REGION Network 10: Concatenadora 10
   RUNG wire#powerrail
      Contact( "EstadosCmpALTA-MTA"._6s1 )
      I_Contact( "CompALTA-MTA".ReqMch6 )
      wire#w1
      Contact( "DB-CompAltaDatos".Aut6 )
      Coil( "Concatenadoras"._6c10 )
   END_RUNG
   RUNG wire#powerrail
      Contact( "EstadosCmpALTA-MTA"._6s9 )
      I_Contact( "CompALTA-MTA".ReqMch6 )
   END_RUNG wire#w1
   RUNG wire#powerrail
      Contact( "EstadosCmpALTA-MTA"._6s3 )
      I_Contact( "DB-CompAltaDatos".PanMchCmp6 )
   END_RUNG wire#w1
   // the same network as SCL:
   "Concatenadoras"._6c10 := (("EstadosCmpALTA-MTA"._6s1 AND NOT "CompALTA-MTA".ReqMch6) OR ("EstadosCmpALTA-MTA"._6s9 AND NOT "CompALTA-MTA".ReqMch6) OR ("EstadosCmpALTA-MTA"._6s3 AND NOT "DB-CompAltaDatos".PanMchCmp6)) AND "DB-CompAltaDatos".Aut6;
END_REGION

REGION Network 11: Concatenadora 4
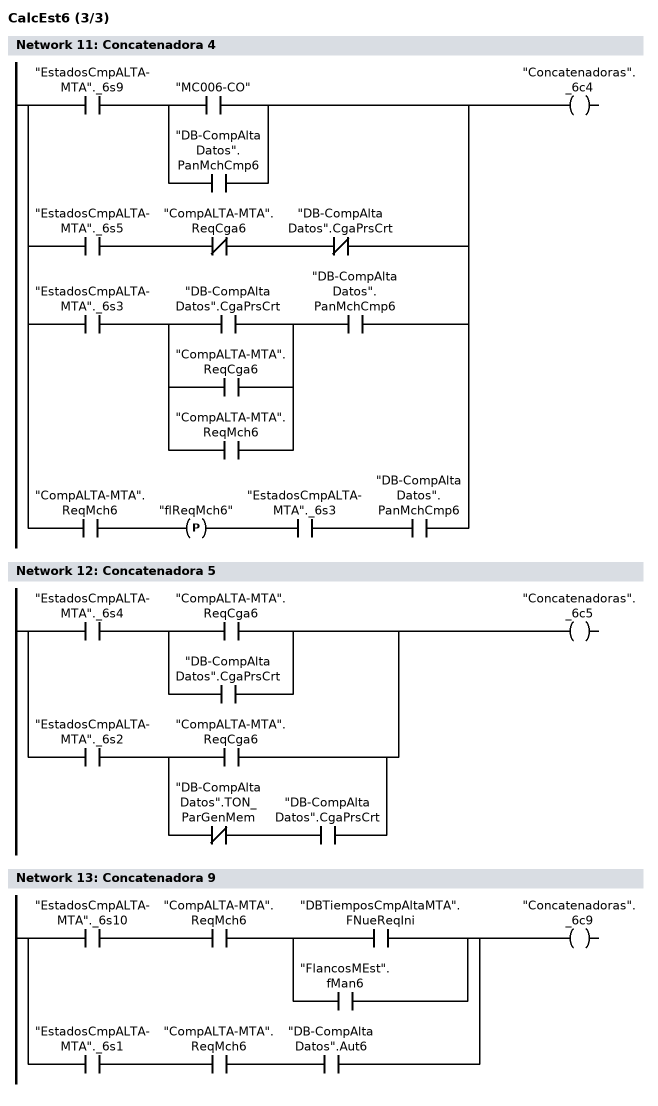
   RUNG wire#powerrail
      Contact( "EstadosCmpALTA-MTA"._6s9 )
      wire#w1
      Contact( "MC006-CO" )
      wire#w2
      Coil( "Concatenadoras"._6c4 )
   END_RUNG
   RUNG wire#w1
      Contact( "DB-CompAltaDatos".PanMchCmp6 )
   END_RUNG wire#w2
   RUNG wire#powerrail
      Contact( "EstadosCmpALTA-MTA"._6s5 )
      I_Contact( "CompALTA-MTA".ReqCga6 )
      I_Contact( "DB-CompAltaDatos".CgaPrsCrt )
   END_RUNG wire#w2
   RUNG wire#powerrail
      Contact( "EstadosCmpALTA-MTA"._6s3 )
      wire#w3
      Contact( "DB-CompAltaDatos".CgaPrsCrt )
      wire#w4
      Contact( "DB-CompAltaDatos".PanMchCmp6 )
   END_RUNG wire#w2
   RUNG wire#w3
      Contact( "CompALTA-MTA".ReqCga6 )
   END_RUNG wire#w4
   RUNG wire#w3
      Contact( "CompALTA-MTA".ReqMch6 )
   END_RUNG wire#w4
   RUNG wire#powerrail
      Contact( "CompALTA-MTA".ReqMch6 )
      P_Trig( "flReqMch6" )
      Contact( "EstadosCmpALTA-MTA"._6s3 )
      Contact( "DB-CompAltaDatos".PanMchCmp6 )
   END_RUNG wire#w2
   // the same network as SCL:
   #_w1 := "CompALTA-MTA".ReqMch6 AND NOT "flReqMch6";   // rising edge
   "flReqMch6" := "CompALTA-MTA".ReqMch6;
   "Concatenadoras"._6c4 := ("EstadosCmpALTA-MTA"._6s9 AND ("MC006-CO" OR "DB-CompAltaDatos".PanMchCmp6)) OR ("EstadosCmpALTA-MTA"._6s5 AND NOT "CompALTA-MTA".ReqCga6 AND NOT "DB-CompAltaDatos".CgaPrsCrt) OR ("EstadosCmpALTA-MTA"._6s3 AND ("DB-CompAltaDatos".CgaPrsCrt OR "CompALTA-MTA".ReqCga6 OR "CompALTA-MTA".ReqMch6) AND "DB-CompAltaDatos".PanMchCmp6) OR (#_w1 AND "EstadosCmpALTA-MTA"._6s3 AND "DB-CompAltaDatos".PanMchCmp6);
END_REGION

REGION Network 12: Concatenadora 5
   RUNG wire#powerrail
      Contact( "EstadosCmpALTA-MTA"._6s4 )
      wire#w1
      Contact( "CompALTA-MTA".ReqCga6 )
      wire#w2
      Coil( "Concatenadoras"._6c5 )
   END_RUNG
   RUNG wire#w1
      Contact( "DB-CompAltaDatos".CgaPrsCrt )
   END_RUNG wire#w2
   RUNG wire#powerrail
      Contact( "EstadosCmpALTA-MTA"._6s2 )
      wire#w3
      Contact( "CompALTA-MTA".ReqCga6 )
   END_RUNG wire#w2
   RUNG wire#w3
      I_Contact( "DB-CompAltaDatos".TON_ParGenMem )
      Contact( "DB-CompAltaDatos".CgaPrsCrt )
   END_RUNG wire#w2
   // the same network as SCL:
   "Concatenadoras"._6c5 := ("EstadosCmpALTA-MTA"._6s4 AND ("CompALTA-MTA".ReqCga6 OR "DB-CompAltaDatos".CgaPrsCrt)) OR ("EstadosCmpALTA-MTA"._6s2 AND ("CompALTA-MTA".ReqCga6 OR (NOT "DB-CompAltaDatos".TON_ParGenMem AND "DB-CompAltaDatos".CgaPrsCrt)));
END_REGION

REGION Network 13: Concatenadora 9
   RUNG wire#powerrail
      Contact( "EstadosCmpALTA-MTA"._6s10 )
      Contact( "CompALTA-MTA".ReqMch6 )
      wire#w1
      Contact( "DBTiemposCmpAltaMTA".FNueReqIni )
      wire#w2
      Coil( "Concatenadoras"._6c9 )
   END_RUNG
   RUNG wire#w1
      Contact( "FlancosMEst".fMan6 )
   END_RUNG wire#w2
   RUNG wire#powerrail
      Contact( "EstadosCmpALTA-MTA"._6s1 )
      Contact( "CompALTA-MTA".ReqMch6 )
      Contact( "DB-CompAltaDatos".Aut6 )
   END_RUNG wire#w2
   // the same network as SCL:
   "Concatenadoras"._6c9 := ("EstadosCmpALTA-MTA"._6s10 AND "CompALTA-MTA".ReqMch6 AND ("DBTiemposCmpAltaMTA".FNueReqIni OR "FlancosMEst".fMan6)) OR ("EstadosCmpALTA-MTA"._6s1 AND "CompALTA-MTA".ReqMch6 AND "DB-CompAltaDatos".Aut6);
END_REGION

REGION Network 14 (STL): Maquina de estados
         CALL  "FC_MAQ_EST_16"
         ( IN0  := %DB127.DBW10,
           IN1  := %DB128.DBW10,
           OUT2 := "ErrPMQ6",
           OUT3 := "ErrCMQ6",
           IO4  := %DB120.DBW10
         );
         NOP   0;
END_REGION

REGION Network 15 (STL): Bloque animación compresor
         CALL  "FC-ANIM-CMP"
         ( IN0  := %DB120.DBW10,
           OUT1 := "CompALTA-MTA".AnimCMP6
         );

         NOP   0;
END_REGION
END_FUNCTION

// folder: Compresores/Baja

FUNCTION "AutoCmpBaja" : Void   // FC24, LAD
{ S7_Optimized_Access := 'FALSE' }
VERSION : 0.1
   VAR_TEMP   // added for the SCL form of the ladder/FBD networks
      _w1 : Bool;
      _s5time1 : S5Time;
      _w2 : Bool;
   END_VAR
BEGIN

REGION Network 1 (STL)
         A(;
         L     "CmpBajaAuto".SPoffMC060;
         L     "CmpBajaAuto".SPonMC060;
         <=R;
         );
         JNB   M001;
         L     "CmpBajaAuto".SPonMC060;
         L     1;
         +R;
         T     "CmpBajaAuto".SPoffMC060;
   M001: NOP   0;
END_REGION

REGION Network 2 (STL)
         A(;
         L     "CmpBajaAuto".SPoffMC061;
         L     "CmpBajaAuto".SPonMC061;
         <=R;
         );
         JNB   M002;
         L     "CmpBajaAuto".SPonMC061;
         L     1;
         +R;
         T     "CmpBajaAuto".SPoffMC061;
   M002: NOP   0;
END_REGION

REGION Network 3 (STL)
         A(;
         L     "CmpBajaAuto".SPoffMC062;
         L     "CmpBajaAuto".SPonMC062;
         <=R;
         );
         JNB   M003;
         L     "CmpBajaAuto".SPonMC062;
         L     1;
         +R;
         T     "CmpBajaAuto".SPoffMC062;
   M003: NOP   0;
END_REGION

REGION Network 4 (STL)
         A(;
         L     "CmpBajaAuto".SPoffMC063;
         L     "CmpBajaAuto".SPonMC063;
         <=R;
         );
         JNB   M004;
         L     "CmpBajaAuto".SPonMC063;
         L     1;
         +R;
         T     "CmpBajaAuto".SPoffMC063;
   M004: NOP   0;
END_REGION

REGION Network 5 (STL)
         A(;
         L     "CmpBajaAuto".SPoffMC064;
         L     "CmpBajaAuto".SPonMC064;
         <=R;
         );
         JNB   M005;
         L     "CmpBajaAuto".SPonMC064;
         L     1;
         +R;
         T     "CmpBajaAuto".SPoffMC064;
   M005: NOP   0;
END_REGION

REGION Network 6
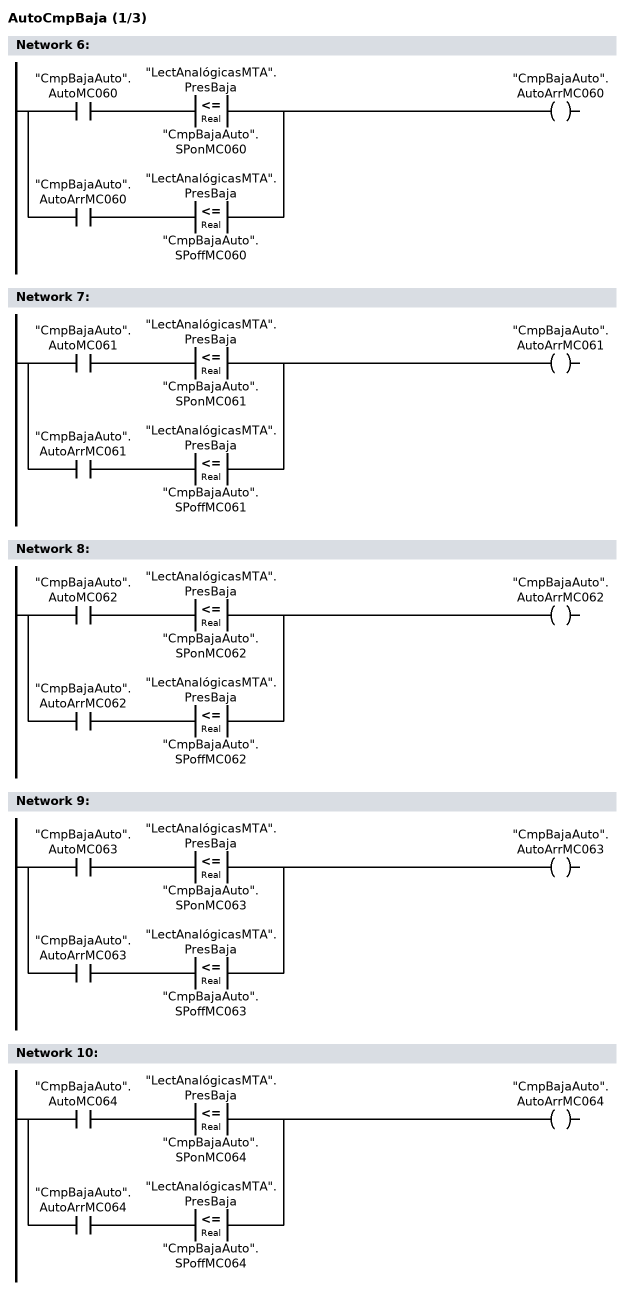
   "CmpBajaAuto".AutoArrMC060 := ("CmpBajaAuto".AutoMC060 AND ("LectAnalógicasMTA".PresBaja <= "CmpBajaAuto".SPonMC060)) OR ("CmpBajaAuto".AutoArrMC060 AND ("LectAnalógicasMTA".PresBaja <= "CmpBajaAuto".SPoffMC060));
END_REGION

REGION Network 7
   "CmpBajaAuto".AutoArrMC061 := ("CmpBajaAuto".AutoMC061 AND ("LectAnalógicasMTA".PresBaja <= "CmpBajaAuto".SPonMC061)) OR ("CmpBajaAuto".AutoArrMC061 AND ("LectAnalógicasMTA".PresBaja <= "CmpBajaAuto".SPoffMC061));
END_REGION

REGION Network 8
   "CmpBajaAuto".AutoArrMC062 := ("CmpBajaAuto".AutoMC062 AND ("LectAnalógicasMTA".PresBaja <= "CmpBajaAuto".SPonMC062)) OR ("CmpBajaAuto".AutoArrMC062 AND ("LectAnalógicasMTA".PresBaja <= "CmpBajaAuto".SPoffMC062));
END_REGION

REGION Network 9
   "CmpBajaAuto".AutoArrMC063 := ("CmpBajaAuto".AutoMC063 AND ("LectAnalógicasMTA".PresBaja <= "CmpBajaAuto".SPonMC063)) OR ("CmpBajaAuto".AutoArrMC063 AND ("LectAnalógicasMTA".PresBaja <= "CmpBajaAuto".SPoffMC063));
END_REGION

REGION Network 10
   "CmpBajaAuto".AutoArrMC064 := ("CmpBajaAuto".AutoMC064 AND ("LectAnalógicasMTA".PresBaja <= "CmpBajaAuto".SPonMC064)) OR ("CmpBajaAuto".AutoArrMC064 AND ("LectAnalógicasMTA".PresBaja <= "CmpBajaAuto".SPoffMC064));
END_REGION

REGION Network 11
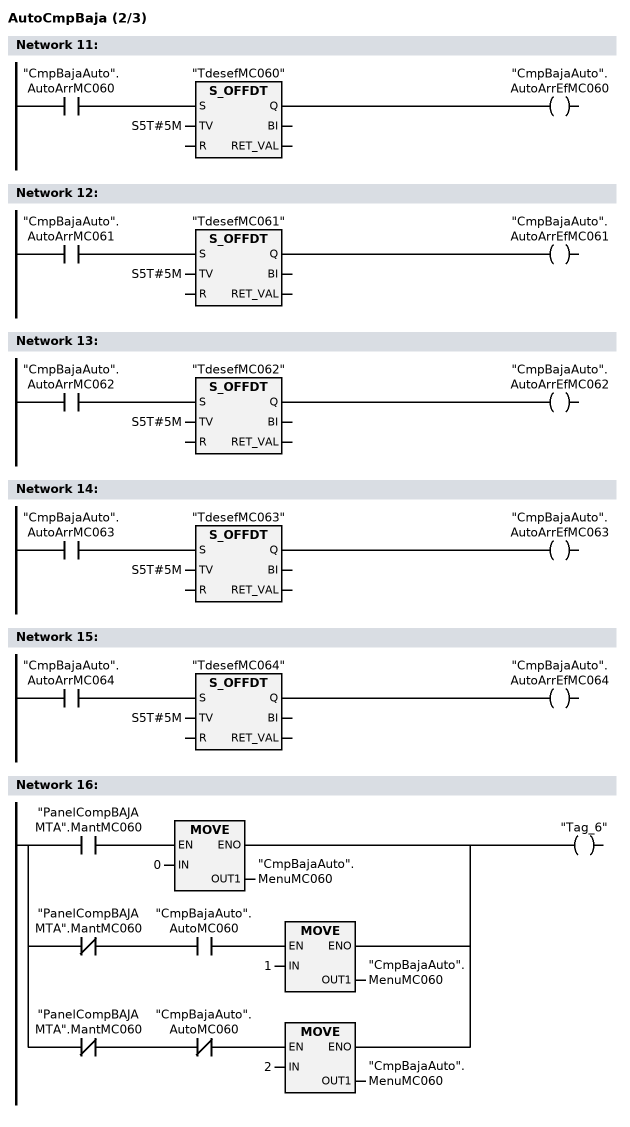
   RUNG wire#powerrail
      Contact( "CmpBajaAuto".AutoArrMC060 )
      S_OFFDT(T_NO := "TdesefMC060", TV := S5T#5M, R :=, BI =>, RET_VAL =>)
      Coil( "CmpBajaAuto".AutoArrEfMC060 )
   END_RUNG
   // the same network as SCL:
   #_s5time1 := S_OFFDT(T_NO := "TdesefMC060", TV := S5T#5M, S := "CmpBajaAuto".AutoArrMC060, Q => #_w1);
   "CmpBajaAuto".AutoArrEfMC060 := #_w1;
END_REGION

REGION Network 12
   RUNG wire#powerrail
      Contact( "CmpBajaAuto".AutoArrMC061 )
      S_OFFDT(T_NO := "TdesefMC061", TV := S5T#5M, R :=, BI =>, RET_VAL =>)
      Coil( "CmpBajaAuto".AutoArrEfMC061 )
   END_RUNG
   // the same network as SCL:
   #_s5time1 := S_OFFDT(T_NO := "TdesefMC061", TV := S5T#5M, S := "CmpBajaAuto".AutoArrMC061, Q => #_w1);
   "CmpBajaAuto".AutoArrEfMC061 := #_w1;
END_REGION

REGION Network 13
   RUNG wire#powerrail
      Contact( "CmpBajaAuto".AutoArrMC062 )
      S_OFFDT(T_NO := "TdesefMC062", TV := S5T#5M, R :=, BI =>, RET_VAL =>)
      Coil( "CmpBajaAuto".AutoArrEfMC062 )
   END_RUNG
   // the same network as SCL:
   #_s5time1 := S_OFFDT(T_NO := "TdesefMC062", TV := S5T#5M, S := "CmpBajaAuto".AutoArrMC062, Q => #_w1);
   "CmpBajaAuto".AutoArrEfMC062 := #_w1;
END_REGION

REGION Network 14
   RUNG wire#powerrail
      Contact( "CmpBajaAuto".AutoArrMC063 )
      S_OFFDT(T_NO := "TdesefMC063", TV := S5T#5M, R :=, BI =>, RET_VAL =>)
      Coil( "CmpBajaAuto".AutoArrEfMC063 )
   END_RUNG
   // the same network as SCL:
   #_s5time1 := S_OFFDT(T_NO := "TdesefMC063", TV := S5T#5M, S := "CmpBajaAuto".AutoArrMC063, Q => #_w1);
   "CmpBajaAuto".AutoArrEfMC063 := #_w1;
END_REGION

REGION Network 15
   RUNG wire#powerrail
      Contact( "CmpBajaAuto".AutoArrMC064 )
      S_OFFDT(T_NO := "TdesefMC064", TV := S5T#5M, R :=, BI =>, RET_VAL =>)
      Coil( "CmpBajaAuto".AutoArrEfMC064 )
   END_RUNG
   // the same network as SCL:
   #_s5time1 := S_OFFDT(T_NO := "TdesefMC064", TV := S5T#5M, S := "CmpBajaAuto".AutoArrMC064, Q => #_w1);
   "CmpBajaAuto".AutoArrEfMC064 := #_w1;
END_REGION

REGION Network 16
   RUNG wire#powerrail
      Contact( "PanelCompBAJA MTA".MantMC060 )
      { S7_GenerateENO := "TRUE" } Move(in := 0, out1 => "CmpBajaAuto".MenuMC060)
      wire#w1
      Coil( "Tag_6" )
   END_RUNG
   RUNG wire#powerrail
      I_Contact( "PanelCompBAJA MTA".MantMC060 )
      Contact( "CmpBajaAuto".AutoMC060 )
      { S7_GenerateENO := "TRUE" } Move(in := 1, out1 => "CmpBajaAuto".MenuMC060)
   END_RUNG wire#w1
   RUNG wire#powerrail
      I_Contact( "PanelCompBAJA MTA".MantMC060 )
      I_Contact( "CmpBajaAuto".AutoMC060 )
      { S7_GenerateENO := "TRUE" } Move(in := 2, out1 => "CmpBajaAuto".MenuMC060)
   END_RUNG wire#w1
   // the same network as SCL:
   // ENO of a box is taken as its EN; it also drops when the box reports an error
   IF "PanelCompBAJA MTA".MantMC060 THEN "CmpBajaAuto".MenuMC060 := 0; END_IF;
   #_w1 := NOT "PanelCompBAJA MTA".MantMC060 AND "CmpBajaAuto".AutoMC060;
   IF #_w1 THEN "CmpBajaAuto".MenuMC060 := 1; END_IF;
   #_w2 := NOT "PanelCompBAJA MTA".MantMC060 AND NOT "CmpBajaAuto".AutoMC060;
   IF #_w2 THEN "CmpBajaAuto".MenuMC060 := 2; END_IF;
   "Tag_6" := "PanelCompBAJA MTA".MantMC060 OR #_w1 OR #_w2;
END_REGION

REGION Network 17
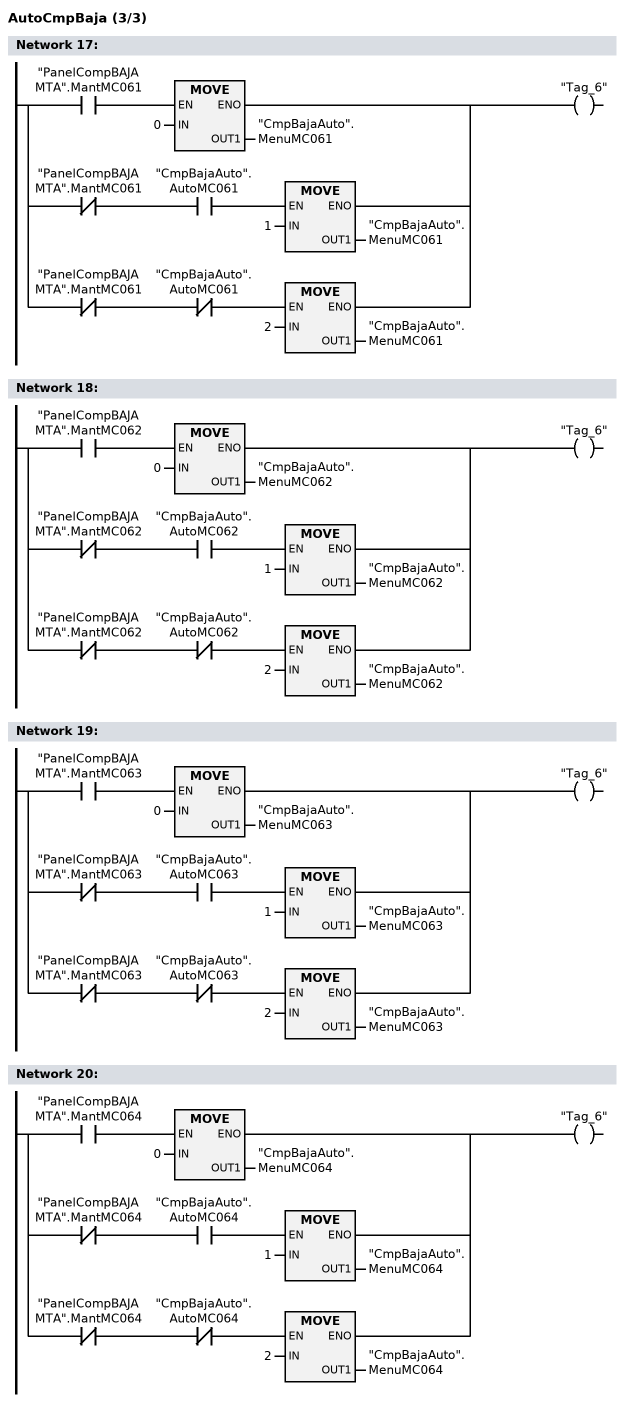
   RUNG wire#powerrail
      Contact( "PanelCompBAJA MTA".MantMC061 )
      { S7_GenerateENO := "TRUE" } Move(in := 0, out1 => "CmpBajaAuto".MenuMC061)
      wire#w1
      Coil( "Tag_6" )
   END_RUNG
   RUNG wire#powerrail
      I_Contact( "PanelCompBAJA MTA".MantMC061 )
      Contact( "CmpBajaAuto".AutoMC061 )
      { S7_GenerateENO := "TRUE" } Move(in := 1, out1 => "CmpBajaAuto".MenuMC061)
   END_RUNG wire#w1
   RUNG wire#powerrail
      I_Contact( "PanelCompBAJA MTA".MantMC061 )
      I_Contact( "CmpBajaAuto".AutoMC061 )
      { S7_GenerateENO := "TRUE" } Move(in := 2, out1 => "CmpBajaAuto".MenuMC061)
   END_RUNG wire#w1
   // the same network as SCL:
   // ENO of a box is taken as its EN; it also drops when the box reports an error
   IF "PanelCompBAJA MTA".MantMC061 THEN "CmpBajaAuto".MenuMC061 := 0; END_IF;
   #_w1 := NOT "PanelCompBAJA MTA".MantMC061 AND "CmpBajaAuto".AutoMC061;
   IF #_w1 THEN "CmpBajaAuto".MenuMC061 := 1; END_IF;
   #_w2 := NOT "PanelCompBAJA MTA".MantMC061 AND NOT "CmpBajaAuto".AutoMC061;
   IF #_w2 THEN "CmpBajaAuto".MenuMC061 := 2; END_IF;
   "Tag_6" := "PanelCompBAJA MTA".MantMC061 OR #_w1 OR #_w2;
END_REGION

REGION Network 18
   RUNG wire#powerrail
      Contact( "PanelCompBAJA MTA".MantMC062 )
      { S7_GenerateENO := "TRUE" } Move(in := 0, out1 => "CmpBajaAuto".MenuMC062)
      wire#w1
      Coil( "Tag_6" )
   END_RUNG
   RUNG wire#powerrail
      I_Contact( "PanelCompBAJA MTA".MantMC062 )
      Contact( "CmpBajaAuto".AutoMC062 )
      { S7_GenerateENO := "TRUE" } Move(in := 1, out1 => "CmpBajaAuto".MenuMC062)
   END_RUNG wire#w1
   RUNG wire#powerrail
      I_Contact( "PanelCompBAJA MTA".MantMC062 )
      I_Contact( "CmpBajaAuto".AutoMC062 )
      { S7_GenerateENO := "TRUE" } Move(in := 2, out1 => "CmpBajaAuto".MenuMC062)
   END_RUNG wire#w1
   // the same network as SCL:
   // ENO of a box is taken as its EN; it also drops when the box reports an error
   IF "PanelCompBAJA MTA".MantMC062 THEN "CmpBajaAuto".MenuMC062 := 0; END_IF;
   #_w1 := NOT "PanelCompBAJA MTA".MantMC062 AND "CmpBajaAuto".AutoMC062;
   IF #_w1 THEN "CmpBajaAuto".MenuMC062 := 1; END_IF;
   #_w2 := NOT "PanelCompBAJA MTA".MantMC062 AND NOT "CmpBajaAuto".AutoMC062;
   IF #_w2 THEN "CmpBajaAuto".MenuMC062 := 2; END_IF;
   "Tag_6" := "PanelCompBAJA MTA".MantMC062 OR #_w1 OR #_w2;
END_REGION

REGION Network 19
   RUNG wire#powerrail
      Contact( "PanelCompBAJA MTA".MantMC063 )
      { S7_GenerateENO := "TRUE" } Move(in := 0, out1 => "CmpBajaAuto".MenuMC063)
      wire#w1
      Coil( "Tag_6" )
   END_RUNG
   RUNG wire#powerrail
      I_Contact( "PanelCompBAJA MTA".MantMC063 )
      Contact( "CmpBajaAuto".AutoMC063 )
      { S7_GenerateENO := "TRUE" } Move(in := 1, out1 => "CmpBajaAuto".MenuMC063)
   END_RUNG wire#w1
   RUNG wire#powerrail
      I_Contact( "PanelCompBAJA MTA".MantMC063 )
      I_Contact( "CmpBajaAuto".AutoMC063 )
      { S7_GenerateENO := "TRUE" } Move(in := 2, out1 => "CmpBajaAuto".MenuMC063)
   END_RUNG wire#w1
   // the same network as SCL:
   // ENO of a box is taken as its EN; it also drops when the box reports an error
   IF "PanelCompBAJA MTA".MantMC063 THEN "CmpBajaAuto".MenuMC063 := 0; END_IF;
   #_w1 := NOT "PanelCompBAJA MTA".MantMC063 AND "CmpBajaAuto".AutoMC063;
   IF #_w1 THEN "CmpBajaAuto".MenuMC063 := 1; END_IF;
   #_w2 := NOT "PanelCompBAJA MTA".MantMC063 AND NOT "CmpBajaAuto".AutoMC063;
   IF #_w2 THEN "CmpBajaAuto".MenuMC063 := 2; END_IF;
   "Tag_6" := "PanelCompBAJA MTA".MantMC063 OR #_w1 OR #_w2;
END_REGION

REGION Network 20
   RUNG wire#powerrail
      Contact( "PanelCompBAJA MTA".MantMC064 )
      { S7_GenerateENO := "TRUE" } Move(in := 0, out1 => "CmpBajaAuto".MenuMC064)
      wire#w1
      Coil( "Tag_6" )
   END_RUNG
   RUNG wire#powerrail
      I_Contact( "PanelCompBAJA MTA".MantMC064 )
      Contact( "CmpBajaAuto".AutoMC064 )
      { S7_GenerateENO := "TRUE" } Move(in := 1, out1 => "CmpBajaAuto".MenuMC064)
   END_RUNG wire#w1
   RUNG wire#powerrail
      I_Contact( "PanelCompBAJA MTA".MantMC064 )
      I_Contact( "CmpBajaAuto".AutoMC064 )
      { S7_GenerateENO := "TRUE" } Move(in := 2, out1 => "CmpBajaAuto".MenuMC064)
   END_RUNG wire#w1
   // the same network as SCL:
   // ENO of a box is taken as its EN; it also drops when the box reports an error
   IF "PanelCompBAJA MTA".MantMC064 THEN "CmpBajaAuto".MenuMC064 := 0; END_IF;
   #_w1 := NOT "PanelCompBAJA MTA".MantMC064 AND "CmpBajaAuto".AutoMC064;
   IF #_w1 THEN "CmpBajaAuto".MenuMC064 := 1; END_IF;
   #_w2 := NOT "PanelCompBAJA MTA".MantMC064 AND NOT "CmpBajaAuto".AutoMC064;
   IF #_w2 THEN "CmpBajaAuto".MenuMC064 := 2; END_IF;
   "Tag_6" := "PanelCompBAJA MTA".MantMC064 OR #_w1 OR #_w2;
END_REGION
END_FUNCTION

// folder: Entradas Analógicas

FUNCTION "LecturasAnalógicasMTA" : Void   // FC15, LAD
{ S7_Optimized_Access := 'FALSE' }
VERSION : 0.1
BEGIN

REGION Network 1: Lectura Temperatura Torres Cavaleto
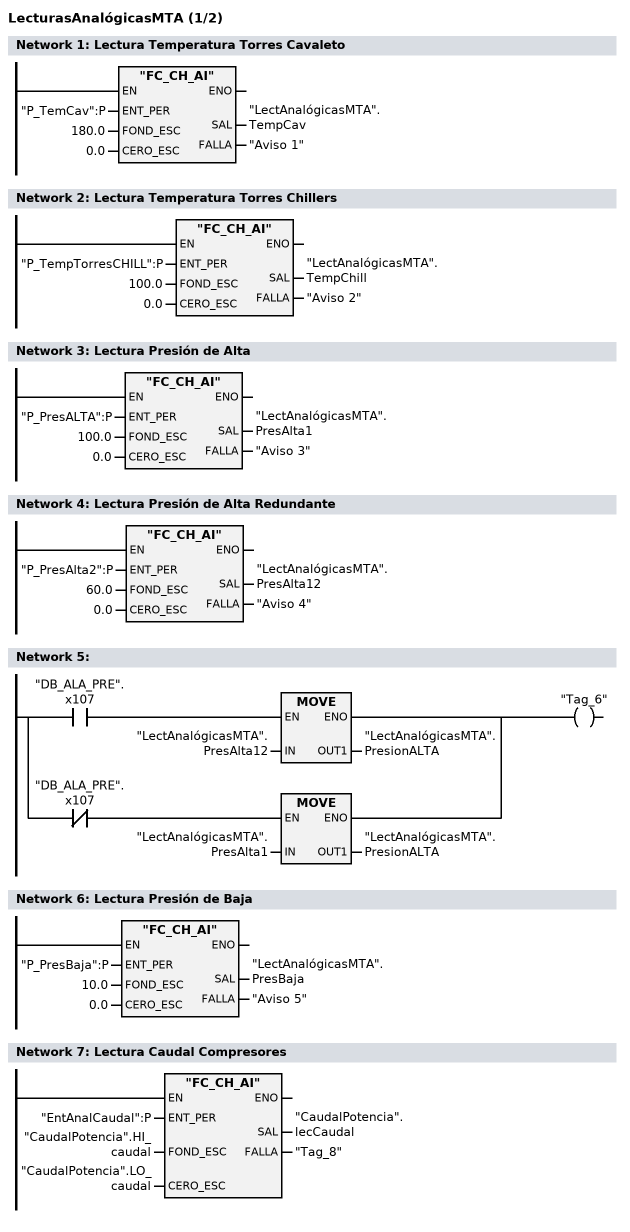
   RUNG wire#powerrail
      "FC_CH_AI"(ENT_PER := "P_TemCav":P, FOND_ESC := 180.0, CERO_ESC := 0.0, SAL => "LectAnalógicasMTA".TempCav, FALLA => "Aviso 1")
   END_RUNG
   // the same network as SCL:
   "FC_CH_AI"(ENT_PER := "P_TemCav":P,
              FOND_ESC := 180.0,
              CERO_ESC := 0.0,
              SAL => "LectAnalógicasMTA".TempCav,
              FALLA => "Aviso 1");
END_REGION

REGION Network 2: Lectura Temperatura Torres Chillers
   RUNG wire#powerrail
      "FC_CH_AI"(ENT_PER := "P_TempTorresCHILL":P, FOND_ESC := 100.0, CERO_ESC := 0.0, SAL => "LectAnalógicasMTA".TempChill, FALLA => "Aviso 2")
   END_RUNG
   // the same network as SCL:
   "FC_CH_AI"(ENT_PER := "P_TempTorresCHILL":P,
              FOND_ESC := 100.0,
              CERO_ESC := 0.0,
              SAL => "LectAnalógicasMTA".TempChill,
              FALLA => "Aviso 2");
END_REGION

REGION Network 3: Lectura Presión de Alta
   RUNG wire#powerrail
      "FC_CH_AI"(ENT_PER := "P_PresALTA":P, FOND_ESC := 100.0, CERO_ESC := 0.0, SAL => "LectAnalógicasMTA".PresAlta1, FALLA => "Aviso 3")
   END_RUNG
   // the same network as SCL:
   "FC_CH_AI"(ENT_PER := "P_PresALTA":P,
              FOND_ESC := 100.0,
              CERO_ESC := 0.0,
              SAL => "LectAnalógicasMTA".PresAlta1,
              FALLA => "Aviso 3");
END_REGION

REGION Network 4: Lectura Presión de Alta Redundante
   RUNG wire#powerrail
      "FC_CH_AI"(ENT_PER := "P_PresAlta2":P, FOND_ESC := 60.0, CERO_ESC := 0.0, SAL => "LectAnalógicasMTA".PresAlta12, FALLA => "Aviso 4")
   END_RUNG
   // the same network as SCL:
   "FC_CH_AI"(ENT_PER := "P_PresAlta2":P,
              FOND_ESC := 60.0,
              CERO_ESC := 0.0,
              SAL => "LectAnalógicasMTA".PresAlta12,
              FALLA => "Aviso 4");
END_REGION

REGION Network 5
   RUNG wire#powerrail
      Contact( "DB_ALA_PRE".x107 )
      { S7_GenerateENO := "TRUE" } Move(in := "LectAnalógicasMTA".PresAlta12, out1 => "LectAnalógicasMTA".PresionALTA)
      wire#w1
      Coil( "Tag_6" )
   END_RUNG
   RUNG wire#powerrail
      I_Contact( "DB_ALA_PRE".x107 )
      { S7_GenerateENO := "TRUE" } Move(in := "LectAnalógicasMTA".PresAlta1, out1 => "LectAnalógicasMTA".PresionALTA)
   END_RUNG wire#w1
   // the same network as SCL:
   // ENO of a box is taken as its EN; it also drops when the box reports an error
   IF "DB_ALA_PRE".x107 THEN "LectAnalógicasMTA".PresionALTA := "LectAnalógicasMTA".PresAlta12; END_IF;
   IF NOT "DB_ALA_PRE".x107 THEN "LectAnalógicasMTA".PresionALTA := "LectAnalógicasMTA".PresAlta1; END_IF;
   "Tag_6" := "DB_ALA_PRE".x107 OR NOT "DB_ALA_PRE".x107;
END_REGION

REGION Network 6: Lectura Presión de Baja
   RUNG wire#powerrail
      "FC_CH_AI"(ENT_PER := "P_PresBaja":P, FOND_ESC := 10.0, CERO_ESC := 0.0, SAL => "LectAnalógicasMTA".PresBaja, FALLA => "Aviso 5")
   END_RUNG
   // the same network as SCL:
   "FC_CH_AI"(ENT_PER := "P_PresBaja":P,
              FOND_ESC := 10.0,
              CERO_ESC := 0.0,
              SAL => "LectAnalógicasMTA".PresBaja,
              FALLA => "Aviso 5");
END_REGION

REGION Network 7: Lectura Caudal Compresores
   RUNG wire#powerrail
      "FC_CH_AI"(ENT_PER := "EntAnalCaudal":P, FOND_ESC := "CaudalPotencia".HI_caudal, CERO_ESC := "CaudalPotencia".LO_caudal, SAL => "CaudalPotencia".lecCaudal, FALLA => "Tag_8")
   END_RUNG
   // the same network as SCL:
   "FC_CH_AI"(ENT_PER := "EntAnalCaudal":P,
              FOND_ESC := "CaudalPotencia".HI_caudal,
              CERO_ESC := "CaudalPotencia".LO_caudal,
              SAL => "CaudalPotencia".lecCaudal,
              FALLA => "Tag_8");
END_REGION

REGION Network 8: Lectura Potencia Compresores
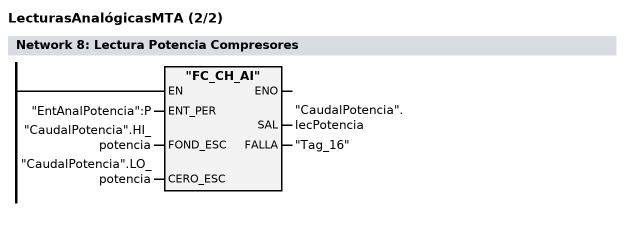
   RUNG wire#powerrail
      "FC_CH_AI"(ENT_PER := "EntAnalPotencia":P, FOND_ESC := "CaudalPotencia".HI_potencia, CERO_ESC := "CaudalPotencia".LO_potencia, SAL => "CaudalPotencia".lecPotencia, FALLA => "Tag_16")
   END_RUNG
   // the same network as SCL:
   "FC_CH_AI"(ENT_PER := "EntAnalPotencia":P,
              FOND_ESC := "CaudalPotencia".HI_potencia,
              CERO_ESC := "CaudalPotencia".LO_potencia,
              SAL => "CaudalPotencia".lecPotencia,
              FALLA => "Tag_16");
END_REGION
END_FUNCTION

// folder: Horas de Marcha

ORGANIZATION_BLOCK "CYC_INT5"   // OB35, LAD
{ S7_Optimized_Access := 'FALSE' }
VERSION : 0.1
   VAR_TEMP   // added for the SCL form of the ladder/FBD networks
      _w1 : Bool;
      _w2 : Bool;
      _w3 : Bool;
      _w4 : Bool;
   END_VAR
BEGIN

REGION Network 1 (STL)
         A     "MC001";
         A     "MC001-CO";
         =     <??.?>;
         A     <??.?>;
         A(;
         L     "SumaOB35 MTA".SMMC001;
         L     600;
         <I;
         );
         JNB   M001;
         L     1;
         L     "SumaOB35 MTA".SMMC001;
         +D;
         T     "SumaOB35 MTA".SMMC001;
   M001: NOP   0;
         A     <??.?>;
         A(;
         L     "SumaOB35 MTA".SMMC001;
         L     600;
         >=I;
         );
         =     <??.?>;
         A     <??.?>;
         JNB   M002;
         L     1;
         L     "SumaOB35 MTA".MMMC001;
         +D;
         T     "SumaOB35 MTA".MMMC001;
   M002: NOP   0;
         A     <??.?>;
         JNB   M003;
         L     0;
         T     "SumaOB35 MTA".SMMC001;
   M003: NOP   0;
         A     <??.?>;
         A(;
         L     "SumaOB35 MTA".MMMC001;
         L     60;
         >=I;
         );
         =     <??.?>;
         A     <??.?>;
         JNB   M004;
         L     1;
         L     "SumaOB35 MTA".HMMC001;
         +D;
         T     "SumaOB35 MTA".HMMC001;
   M004: NOP   0;
         A     <??.?>;
         JNB   M005;
         L     0;
         T     "SumaOB35 MTA".MMMC001;
   M005: NOP   0;
END_REGION

REGION Network 2 (STL)
         A     "MC002";
         A     "MC002-CO";
         =     <??.?>;
         A     <??.?>;
         A(;
         L     "SumaOB35 MTA".SMMC002;
         L     600;
         <I;
         );
         JNB   M006;
         L     1;
         L     "SumaOB35 MTA".SMMC002;
         +D;
         T     "SumaOB35 MTA".SMMC002;
   M006: NOP   0;
         A     <??.?>;
         A(;
         L     "SumaOB35 MTA".SMMC002;
         L     600;
         >=I;
         );
         =     <??.?>;
         A     <??.?>;
         JNB   M007;
         L     1;
         L     "SumaOB35 MTA".MMMC002;
         +D;
         T     "SumaOB35 MTA".MMMC002;
   M007: NOP   0;
         A     <??.?>;
         JNB   M008;
         L     0;
         T     "SumaOB35 MTA".SMMC002;
   M008: NOP   0;
         A     <??.?>;
         A(;
         L     "SumaOB35 MTA".MMMC002;
         L     60;
         >=I;
         );
         =     <??.?>;
         A     <??.?>;
         JNB   M009;
         L     1;
         L     "SumaOB35 MTA".HMMC002;
         +D;
         T     "SumaOB35 MTA".HMMC002;
   M009: NOP   0;
         A     <??.?>;
         JNB   M00a;
         L     0;
         T     "SumaOB35 MTA".MMMC002;
   M00a: NOP   0;
END_REGION

REGION Network 3 (STL)
         A     "MC003";
         A     "MC003-CO";
         =     <??.?>;
         A     <??.?>;
         A(;
         L     "SumaOB35 MTA".SMMC003;
         L     600;
         <I;
         );
         JNB   M00b;
         L     1;
         L     "SumaOB35 MTA".SMMC003;
         +D;
         T     "SumaOB35 MTA".SMMC003;
   M00b: NOP   0;
         A     <??.?>;
         A(;
         L     "SumaOB35 MTA".SMMC003;
         L     600;
         >=I;
         );
         =     <??.?>;
         A     <??.?>;
         JNB   M00c;
         L     1;
         L     "SumaOB35 MTA".MMMC003;
         +D;
         T     "SumaOB35 MTA".MMMC003;
   M00c: NOP   0;
         A     <??.?>;
         JNB   M00d;
         L     0;
         T     "SumaOB35 MTA".SMMC003;
   M00d: NOP   0;
         A     <??.?>;
         A(;
         L     "SumaOB35 MTA".MMMC003;
         L     60;
         >=I;
         );
         =     <??.?>;
         A     <??.?>;
         JNB   M00e;
         L     1;
         L     "SumaOB35 MTA".HMMC003;
         +D;
         T     "SumaOB35 MTA".HMMC003;
   M00e: NOP   0;
         A     <??.?>;
         JNB   M00f;
         L     0;
         T     "SumaOB35 MTA".MMMC003;
   M00f: NOP   0;
END_REGION

REGION Network 4 (STL)
         A     "MC004";
         A     "MC004-CO";
         =     <??.?>;
         A     <??.?>;
         A(;
         L     "SumaOB35 MTA".SMMC004;
         L     600;
         <I;
         );
         JNB   M010;
         L     1;
         L     "SumaOB35 MTA".SMMC004;
         +D;
         T     "SumaOB35 MTA".SMMC004;
   M010: NOP   0;
         A     <??.?>;
         A(;
         L     "SumaOB35 MTA".SMMC004;
         L     600;
         >=I;
         );
         =     <??.?>;
         A     <??.?>;
         JNB   M011;
         L     1;
         L     "SumaOB35 MTA".MMMC004;
         +D;
         T     "SumaOB35 MTA".MMMC004;
   M011: NOP   0;
         A     <??.?>;
         JNB   M012;
         L     0;
         T     "SumaOB35 MTA".SMMC004;
   M012: NOP   0;
         A     <??.?>;
         A(;
         L     "SumaOB35 MTA".MMMC004;
         L     60;
         >=I;
         );
         =     <??.?>;
         A     <??.?>;
         JNB   M013;
         L     1;
         L     "SumaOB35 MTA".HMMC004;
         +D;
         T     "SumaOB35 MTA".HMMC004;
   M013: NOP   0;
         A     <??.?>;
         JNB   M014;
         L     0;
         T     "SumaOB35 MTA".MMMC004;
   M014: NOP   0;
END_REGION

REGION Network 5 (STL)
         A     "MC005";
         A     "MC005-CO";
         =     <??.?>;
         A     <??.?>;
         A(;
         L     "SumaOB35 MTA".SMMC005;
         L     600;
         <I;
         );
         JNB   M015;
         L     1;
         L     "SumaOB35 MTA".SMMC005;
         +D;
         T     "SumaOB35 MTA".SMMC005;
   M015: NOP   0;
         A     <??.?>;
         A(;
         L     "SumaOB35 MTA".SMMC005;
         L     600;
         >=I;
         );
         =     <??.?>;
         A     <??.?>;
         JNB   M016;
         L     1;
         L     "SumaOB35 MTA".MMMC005;
         +D;
         T     "SumaOB35 MTA".MMMC005;
   M016: NOP   0;
         A     <??.?>;
         JNB   M017;
         L     0;
         T     "SumaOB35 MTA".SMMC005;
   M017: NOP   0;
         A     <??.?>;
         A(;
         L     "SumaOB35 MTA".MMMC005;
         L     60;
         >=I;
         );
         =     <??.?>;
         A     <??.?>;
         JNB   M018;
         L     1;
         L     "SumaOB35 MTA".HMMC005;
         +D;
         T     "SumaOB35 MTA".HMMC005;
   M018: NOP   0;
         A     <??.?>;
         JNB   M019;
         L     0;
         T     "SumaOB35 MTA".MMMC005;
   M019: NOP   0;
END_REGION

REGION Network 6 (STL)
         A     "MC006";
         A     "MC006-CO";
         =     <??.?>;
         A     <??.?>;
         A(;
         L     "SumaOB35 MTA".SMMC006;
         L     600;
         <I;
         );
         JNB   M020;
         L     1;
         L     "SumaOB35 MTA".SMMC006;
         +D;
         T     "SumaOB35 MTA".SMMC006;
   M020: NOP   0;
         A     <??.?>;
         A(;
         L     "SumaOB35 MTA".SMMC006;
         L     600;
         >=I;
         );
         =     <??.?>;
         A     <??.?>;
         JNB   M021;
         L     1;
         L     "SumaOB35 MTA".MMMC006;
         +D;
         T     "SumaOB35 MTA".MMMC006;
   M021: NOP   0;
         A     <??.?>;
         JNB   M022;
         L     0;
         T     "SumaOB35 MTA".SMMC006;
   M022: NOP   0;
         A     <??.?>;
         A(;
         L     "SumaOB35 MTA".MMMC006;
         L     60;
         >=I;
         );
         =     <??.?>;
         A     <??.?>;
         JNB   M023;
         L     1;
         L     "SumaOB35 MTA".HMMC006;
         +D;
         T     "SumaOB35 MTA".HMMC006;
   M023: NOP   0;
         A     <??.?>;
         JNB   M024;
         L     0;
         T     "SumaOB35 MTA".MMMC006;
   M024: NOP   0;
END_REGION

REGION Network 7: Encendido de PLC
